(* Logix 5000 project; controller MV vendor 1 type 14 code 217 rev 31.11; software revision 31.00; part 6 of 53 *)
(* tags used below, declared in another part *)
   Alarm_Reset : BOOL;
   Analog_Fault_No : DINT;
   Analog_Simulation_Enabled : BOOL;
   CWD : CHECKWORD_FLAGS;
   Default_Check_Time : DINT;
   FV_YST01_LTX501_AI : PlantItem;   // YST01 LTX501
   FV_YST01_LTX501_AI_RawInput : ALIAS FOR RIO_Rack_2:2:I.Ch2Data;
   FV_YST01_LTX501_ALARM : ALARM_DIGITAL;
   FV_YST01_LTX501_Timer_HiLevel : TIMER;
   FV_YST02_LTX501_AI : PlantItem;   // YST02 LTX501
   FV_YST02_LTX501_AI_RawInput : ALIAS FOR RIO_Rack_2:2:I.Ch3Data;
   FV_YST02_LTX501_ALARM : ALARM_DIGITAL;
   FV_YST02_LTX501_Timer_HiLevel : TIMER;
   FVHRFM03_ALARM : ALARM_DIGITAL;
   FVHRFM03_IP : PlantItem;   // Flow Meter Transmitter
   FVHRFM03_IP_RawInput : ALIAS FOR RIO_Rack_2:16:I.Ch2Data;   // Flow Meter Raw Data
   FVHRLTX02_ALARM : ALARM_DIGITAL;
   FVHRLTX02_IP : PlantItem;   // Effluent Tank Level Transmitter
   FVHRLTX02_IP_Percentage : DINT;
   FVHRLTX02_IP_RawInput : ALIAS FOR RIO_Rack_2:16:I.Ch1Data;   // Effluent Tank Level Transmitter Raw Data
   FVHRLTX02_Timer_HiLevel : TIMER;
   FVHRTM01_IP : PlantItem;   // Turbidty Meter FVHRTM01
   FVHRTM01_IP_RawInput : ALIAS FOR RIO_Rack_2:16:I.Ch0Data;   // Turbidty Meter FVHRTM01 Raw Data
   MC_CH1_CTX1_AI : PlantItem;   // CH1_CTX1
   MC_CH1_CTX1_AI_RawInput : ALIAS FOR RIO_Rack_2:1:I.Ch2Data;   // Real Analog Input , Do Not Use In Code
   MC_CH1_FM_AI : PlantItem;   // CH1_FM
   MC_CH1_FM_AI_RawInput : ALIAS FOR RIO_Rack_2:1:I.Ch4Data;   // Real Analog Input , Do Not Use In Code
   MC_CH1_Log_ID : DINT;
   MC_CH1_PTX_AI : PlantItem;   // CH1_PTX
   MC_CH1_PTX_AI_RawInput : ALIAS FOR RIO_Rack_2:1:I.Ch6Data;   // Real Analog Input , Do Not Use In Code
   MC_CH2_CTX2_AI : PlantItem;   // CH2_CTX2
   MC_CH2_CTX2_AI_RawInput : ALIAS FOR RIO_Rack_2:1:I.Ch3Data;   // Real Analog Input , Do Not Use In Code
   MC_CH2_FM_AI : PlantItem;   // CH2_FM
   MC_CH2_FM_AI_RawInput : ALIAS FOR RIO_Rack_2:1:I.Ch5Data;   // Real Analog Input , Do Not Use In Code
   MC_CH2_Log_ID : DINT;
   MC_CH2_PTX_AI : PlantItem;   // CH2_PTX
   MC_CH2_PTX_AI_RawInput : ALIAS FOR RIO_Rack_2:1:I.Ch7Data;   // Real Analog Input , Do Not Use In Code
   MC_CTX_001_AI : PlantItem;   // CTX_001
   MC_CTX_001_AI_RawInput : ALIAS FOR RIO_Rack_2:1:I.Ch0Data;   // Real Analog Input , Do Not Use In Code
   MC_CTX_002_AI : PlantItem;   // CTX_002
   MC_CTX_002_AI_RawInput : ALIAS FOR RIO_Rack_2:1:I.Ch1Data;   // Real Analog Input , Do Not Use In Code
   MC_N7 : INT[255];   // INTEGER
   MC_P1_SP_AO : PlantItem;   // P1_SP
   MC_P1_SP_AO_RawOutput : ALIAS FOR RIO_Rack_2:3:O.Ch0Data;   // Real Analog Input , Do Not Use In Code
   MC_P2_SP_AO : PlantItem;   // P2_SP
   MC_P2_SP_AO_RawOutput : ALIAS FOR RIO_Rack_2:3:O.Ch1Data;   // Real Analog Input , Do Not Use In Code
   MC_SRV1_Log_ID : DINT;
   MC_SRV2_Log_ID : DINT;
   MC_TTX_001_AI : PlantItem;   // TTX_001
   MC_TTX_001_AI_RawInput : ALIAS FOR RIO_Rack_2:2:I.Ch0Data;   // Real Analog Input , Do Not Use In Code
   MC_TTX_002_AI : PlantItem;   // TTX_002
   MC_TTX_002_AI_RawInput : ALIAS FOR RIO_Rack_2:2:I.Ch1Data;   // Real Analog Input , Do Not Use In Code
   One_Second_One_Scan : ALIAS FOR One_Second_1_scan;
   overrange_RIO_analog_value : REAL;
   underrange_RIO_analog_value : REAL;
   YST_Data : REAL[2];
(* MC_Common, continued *)

ROUTINE MC_A_Events_From_Scada_IDs   (* ladder *)
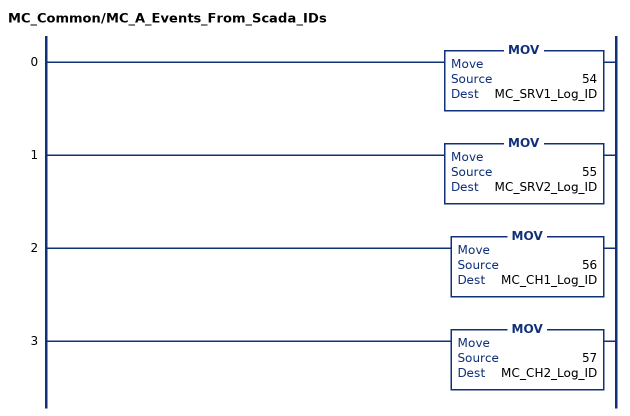
   0: MOV(54,MC_SRV1_Log_ID);
   1: MOV(55,MC_SRV2_Log_ID);
   2: MOV(56,MC_CH1_Log_ID);
   3: MOV(57,MC_CH2_Log_ID);
END_ROUTINE

ROUTINE MC_Analog_Relay_To_NFiles   (* ladder *)
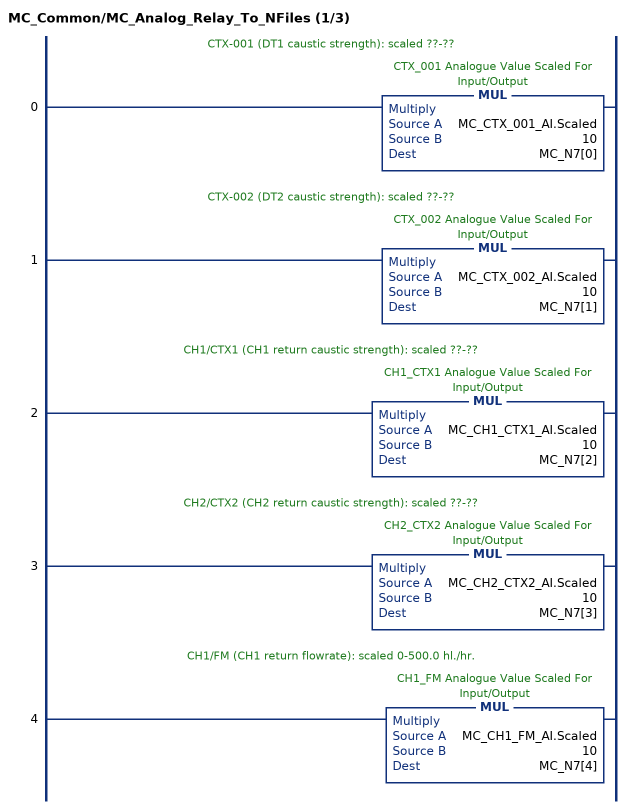
   // CTX-001 (DT1 caustic strength): scaled ??-??
   0: MUL(MC_CTX_001_AI.Scaled,10,MC_N7[0]);
   // CTX-002 (DT2 caustic strength): scaled ??-??
   1: MUL(MC_CTX_002_AI.Scaled,10,MC_N7[1]);
   // CH1/CTX1 (CH1 return caustic strength): scaled ??-??
   2: MUL(MC_CH1_CTX1_AI.Scaled,10,MC_N7[2]);
   // CH2/CTX2 (CH2 return caustic strength): scaled ??-??
   3: MUL(MC_CH2_CTX2_AI.Scaled,10,MC_N7[3]);
   // CH1/FM (CH1 return flowrate): scaled 0-500.0 hl./hr.
   4: MUL(MC_CH1_FM_AI.Scaled,10,MC_N7[4]);
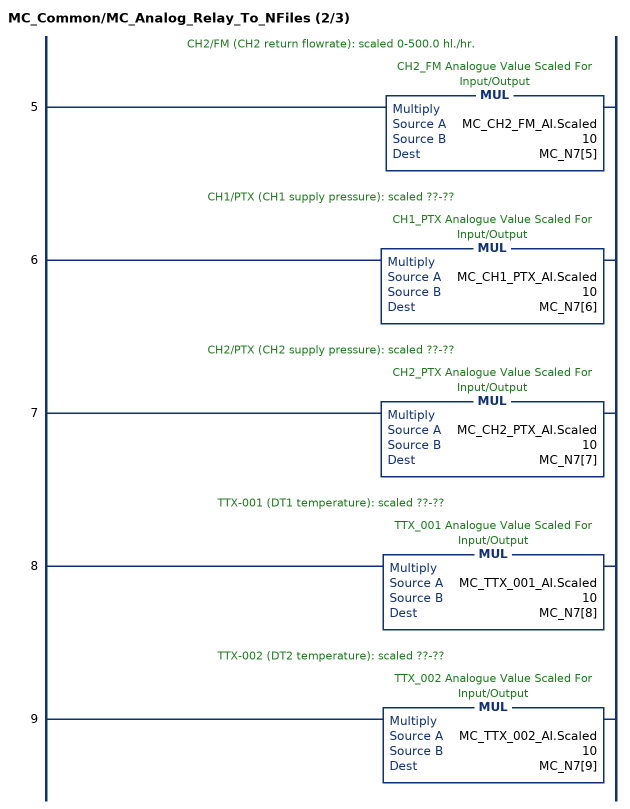
   // CH2/FM (CH2 return flowrate): scaled 0-500.0 hl./hr.
   5: MUL(MC_CH2_FM_AI.Scaled,10,MC_N7[5]);
   // CH1/PTX (CH1 supply pressure): scaled ??-??
   6: MUL(MC_CH1_PTX_AI.Scaled,10,MC_N7[6]);
   // CH2/PTX (CH2 supply pressure): scaled ??-??
   7: MUL(MC_CH2_PTX_AI.Scaled,10,MC_N7[7]);
   // TTX-001 (DT1 temperature): scaled ??-??
   8: MUL(MC_TTX_001_AI.Scaled,10,MC_N7[8]);
   // TTX-002 (DT2 temperature): scaled ??-??
   9: MUL(MC_TTX_002_AI.Scaled,10,MC_N7[9]);
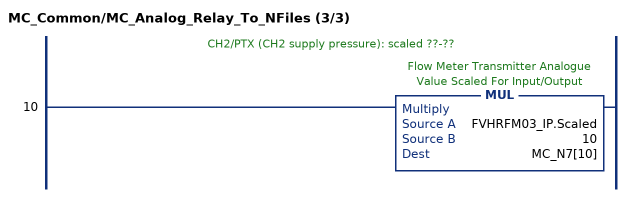
   // CH2/PTX (CH2 supply pressure): scaled ??-??
   10: MUL(FVHRFM03_IP.Scaled,10,MC_N7[10]);
END_ROUTINE

ROUTINE MC_Analogs   (* ladder *)
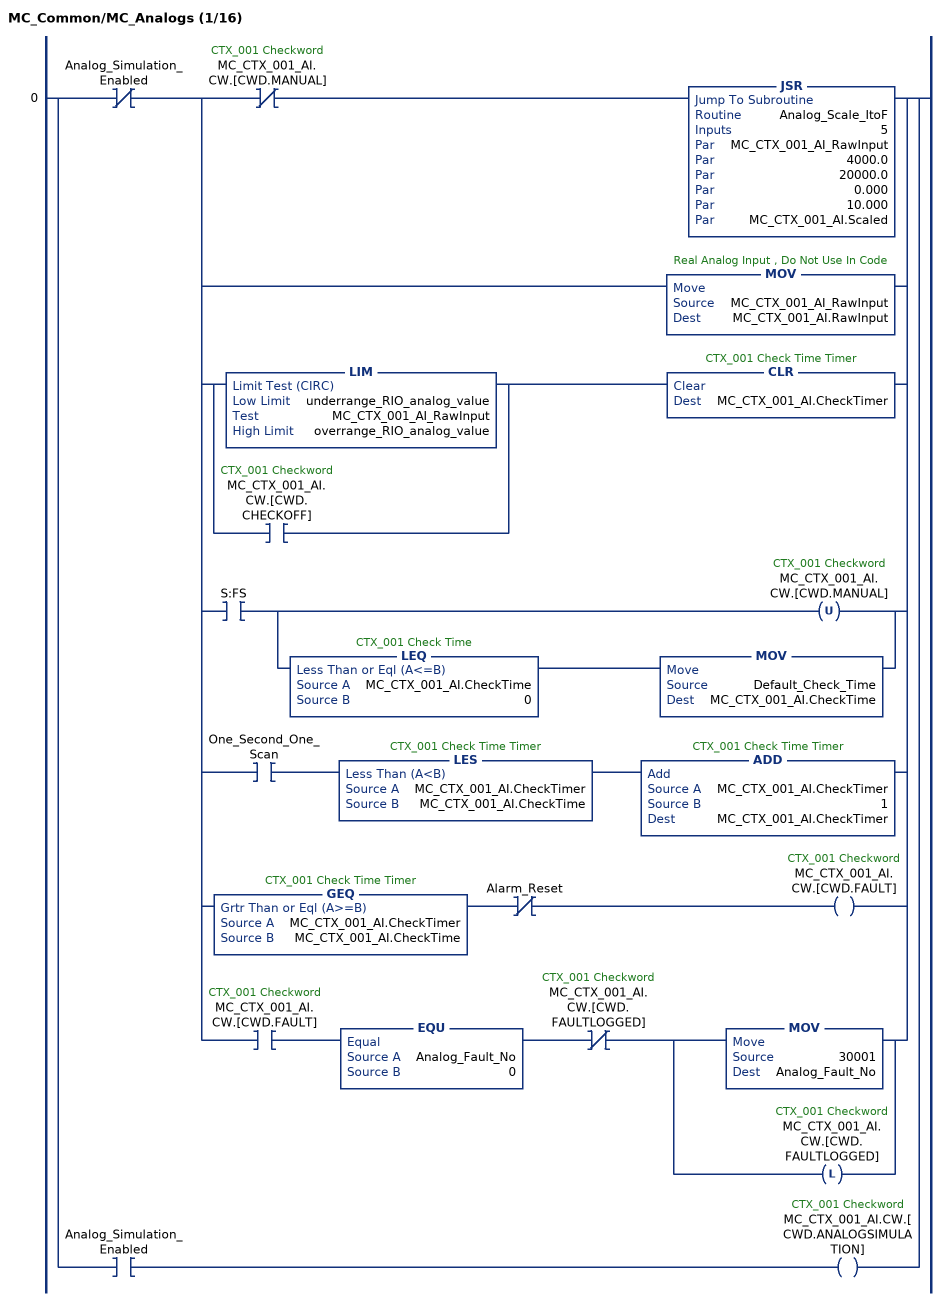
   0: [XIO(Analog_Simulation_Enabled) [XIO(MC_CTX_001_AI.CW.[CWD.MANUAL]) JSR(Analog_Scale_ItoF,5,MC_CTX_001_AI_RawInput,4000.0,20000.0,0.000,10.000,MC_CTX_001_AI.Scaled) ,MOV(MC_CTX_001_AI_RawInput,MC_CTX_001_AI.RawInput) ,[LIM(underrange_RIO_analog_value,MC_CTX_001_AI_RawInput,overrange_RIO_analog_value) ,XIC(MC_CTX_001_AI.CW.[CWD.CHECKOFF]) ] CLR(MC_CTX_001_AI.CheckTimer) ,XIC(S:FS) [OTU(MC_CTX_001_AI.CW.[CWD.MANUAL]) ,LEQ(MC_CTX_001_AI.CheckTime,0) MOV(Default_Check_Time,MC_CTX_001_AI.CheckTime) ] ,XIC(One_Second_One_Scan) LES(MC_CTX_001_AI.CheckTimer,MC_CTX_001_AI.CheckTime) ADD(MC_CTX_001_AI.CheckTimer,1,MC_CTX_001_AI.CheckTimer) ,GEQ(MC_CTX_001_AI.CheckTimer,MC_CTX_001_AI.CheckTime) XIO(Alarm_Reset) OTE(MC_CTX_001_AI.CW.[CWD.FAULT]) ,XIC(MC_CTX_001_AI.CW.[CWD.FAULT]) EQU(Analog_Fault_No,0) XIO(MC_CTX_001_AI.CW.[CWD.FAULTLOGGED]) [MOV(30001,Analog_Fault_No) ,OTL(MC_CTX_001_AI.CW.[CWD.FAULTLOGGED]) ] ] ,XIC(Analog_Simulation_Enabled) OTE(MC_CTX_001_AI.CW.[CWD.ANALOGSIMULATION]) ];
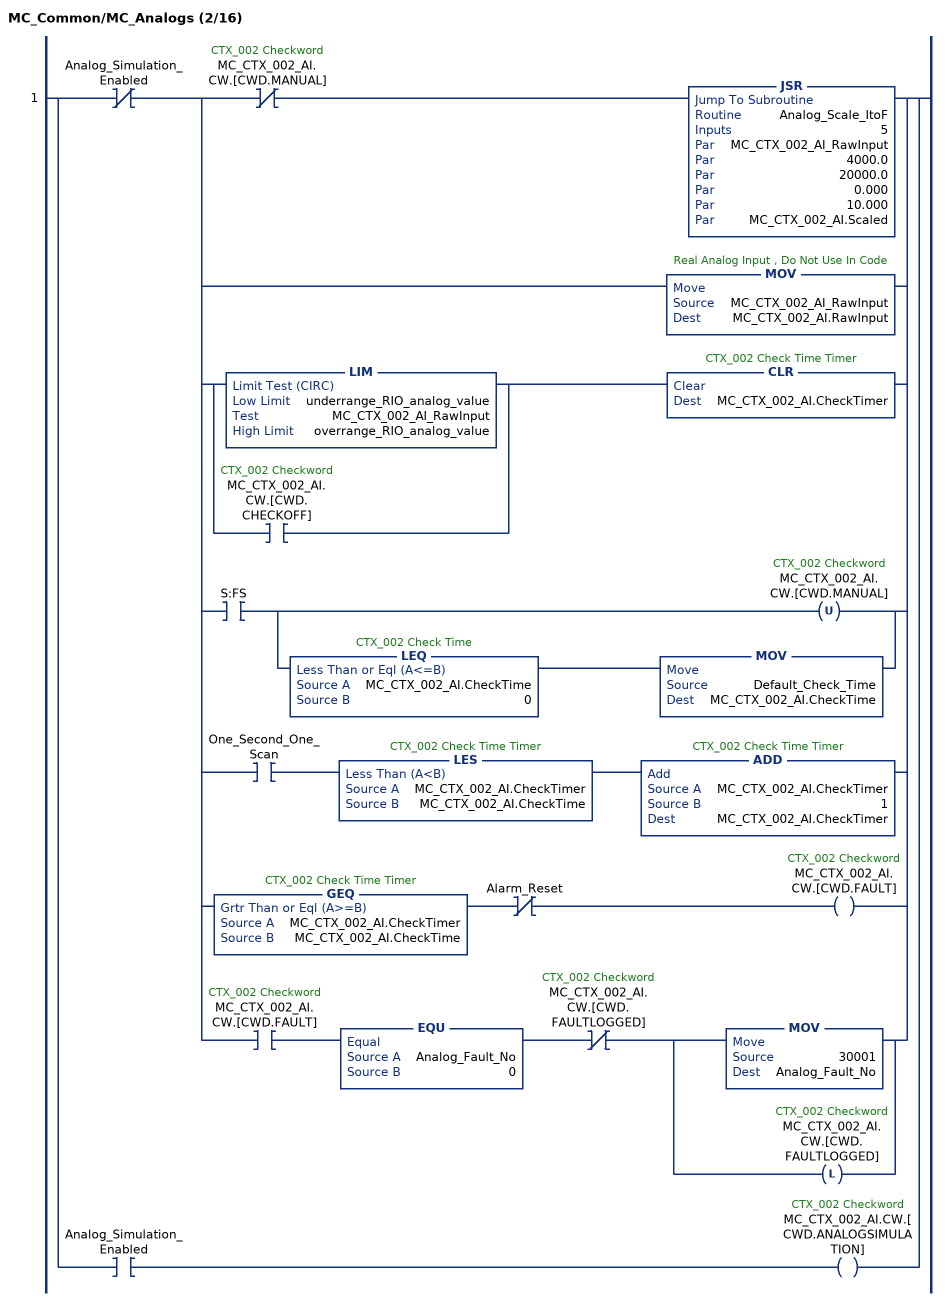
   1: [XIO(Analog_Simulation_Enabled) [XIO(MC_CTX_002_AI.CW.[CWD.MANUAL]) JSR(Analog_Scale_ItoF,5,MC_CTX_002_AI_RawInput,4000.0,20000.0,0.000,10.000,MC_CTX_002_AI.Scaled) ,MOV(MC_CTX_002_AI_RawInput,MC_CTX_002_AI.RawInput) ,[LIM(underrange_RIO_analog_value,MC_CTX_002_AI_RawInput,overrange_RIO_analog_value) ,XIC(MC_CTX_002_AI.CW.[CWD.CHECKOFF]) ] CLR(MC_CTX_002_AI.CheckTimer) ,XIC(S:FS) [OTU(MC_CTX_002_AI.CW.[CWD.MANUAL]) ,LEQ(MC_CTX_002_AI.CheckTime,0) MOV(Default_Check_Time,MC_CTX_002_AI.CheckTime) ] ,XIC(One_Second_One_Scan) LES(MC_CTX_002_AI.CheckTimer,MC_CTX_002_AI.CheckTime) ADD(MC_CTX_002_AI.CheckTimer,1,MC_CTX_002_AI.CheckTimer) ,GEQ(MC_CTX_002_AI.CheckTimer,MC_CTX_002_AI.CheckTime) XIO(Alarm_Reset) OTE(MC_CTX_002_AI.CW.[CWD.FAULT]) ,XIC(MC_CTX_002_AI.CW.[CWD.FAULT]) EQU(Analog_Fault_No,0) XIO(MC_CTX_002_AI.CW.[CWD.FAULTLOGGED]) [MOV(30001,Analog_Fault_No) ,OTL(MC_CTX_002_AI.CW.[CWD.FAULTLOGGED]) ] ] ,XIC(Analog_Simulation_Enabled) OTE(MC_CTX_002_AI.CW.[CWD.ANALOGSIMULATION]) ];
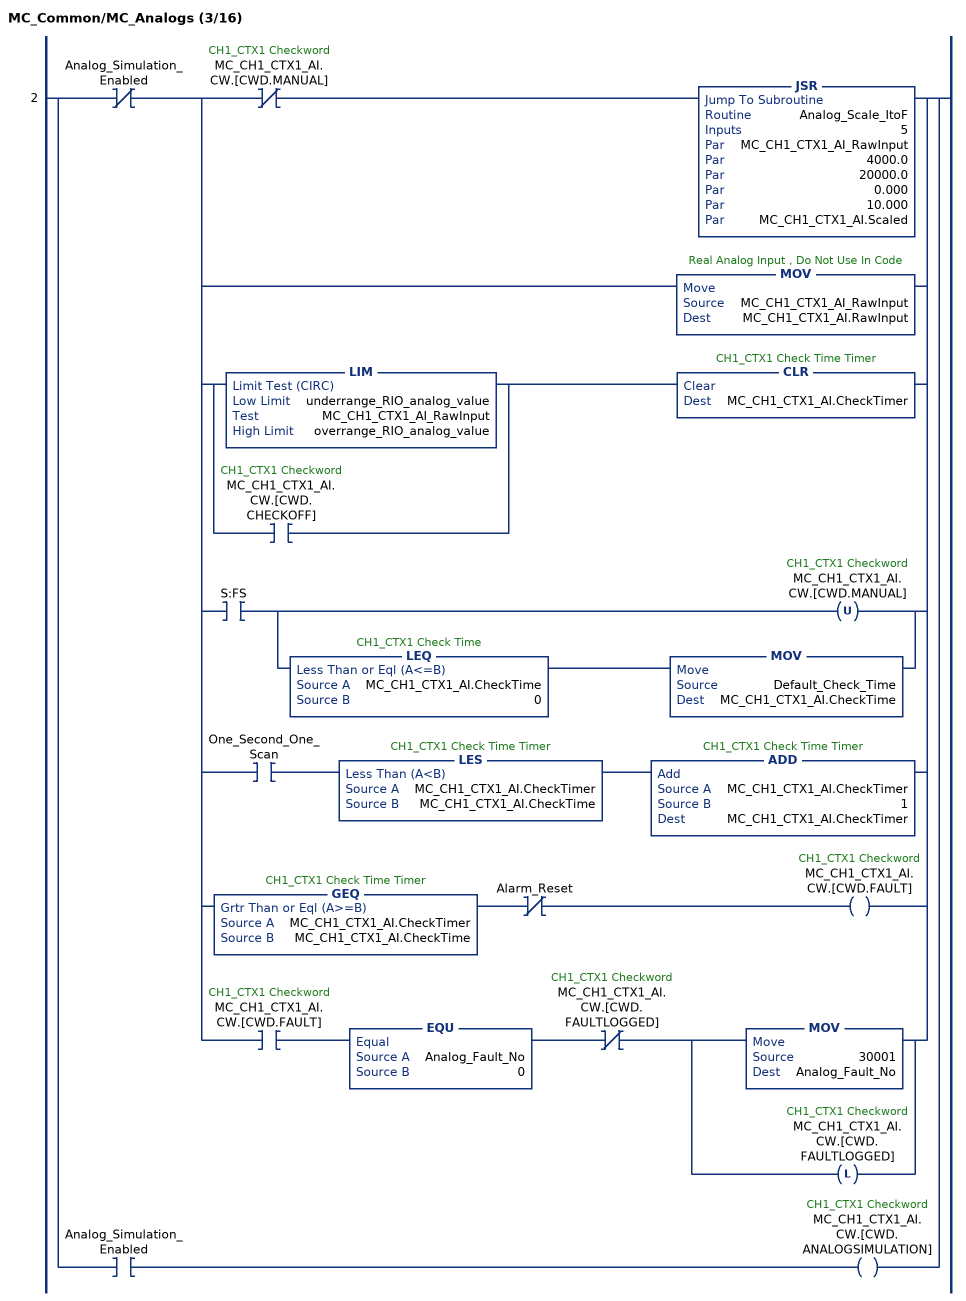
   2: [XIO(Analog_Simulation_Enabled) [XIO(MC_CH1_CTX1_AI.CW.[CWD.MANUAL]) JSR(Analog_Scale_ItoF,5,MC_CH1_CTX1_AI_RawInput,4000.0,20000.0,0.000,10.000,MC_CH1_CTX1_AI.Scaled) ,MOV(MC_CH1_CTX1_AI_RawInput,MC_CH1_CTX1_AI.RawInput) ,[LIM(underrange_RIO_analog_value,MC_CH1_CTX1_AI_RawInput,overrange_RIO_analog_value) ,XIC(MC_CH1_CTX1_AI.CW.[CWD.CHECKOFF]) ] CLR(MC_CH1_CTX1_AI.CheckTimer) ,XIC(S:FS) [OTU(MC_CH1_CTX1_AI.CW.[CWD.MANUAL]) ,LEQ(MC_CH1_CTX1_AI.CheckTime,0) MOV(Default_Check_Time,MC_CH1_CTX1_AI.CheckTime) ] ,XIC(One_Second_One_Scan) LES(MC_CH1_CTX1_AI.CheckTimer,MC_CH1_CTX1_AI.CheckTime) ADD(MC_CH1_CTX1_AI.CheckTimer,1,MC_CH1_CTX1_AI.CheckTimer) ,GEQ(MC_CH1_CTX1_AI.CheckTimer,MC_CH1_CTX1_AI.CheckTime) XIO(Alarm_Reset) OTE(MC_CH1_CTX1_AI.CW.[CWD.FAULT]) ,XIC(MC_CH1_CTX1_AI.CW.[CWD.FAULT]) EQU(Analog_Fault_No,0) XIO(MC_CH1_CTX1_AI.CW.[CWD.FAULTLOGGED]) [MOV(30001,Analog_Fault_No) ,OTL(MC_CH1_CTX1_AI.CW.[CWD.FAULTLOGGED]) ] ] ,XIC(Analog_Simulation_Enabled) OTE(MC_CH1_CTX1_AI.CW.[CWD.ANALOGSIMULATION]) ];
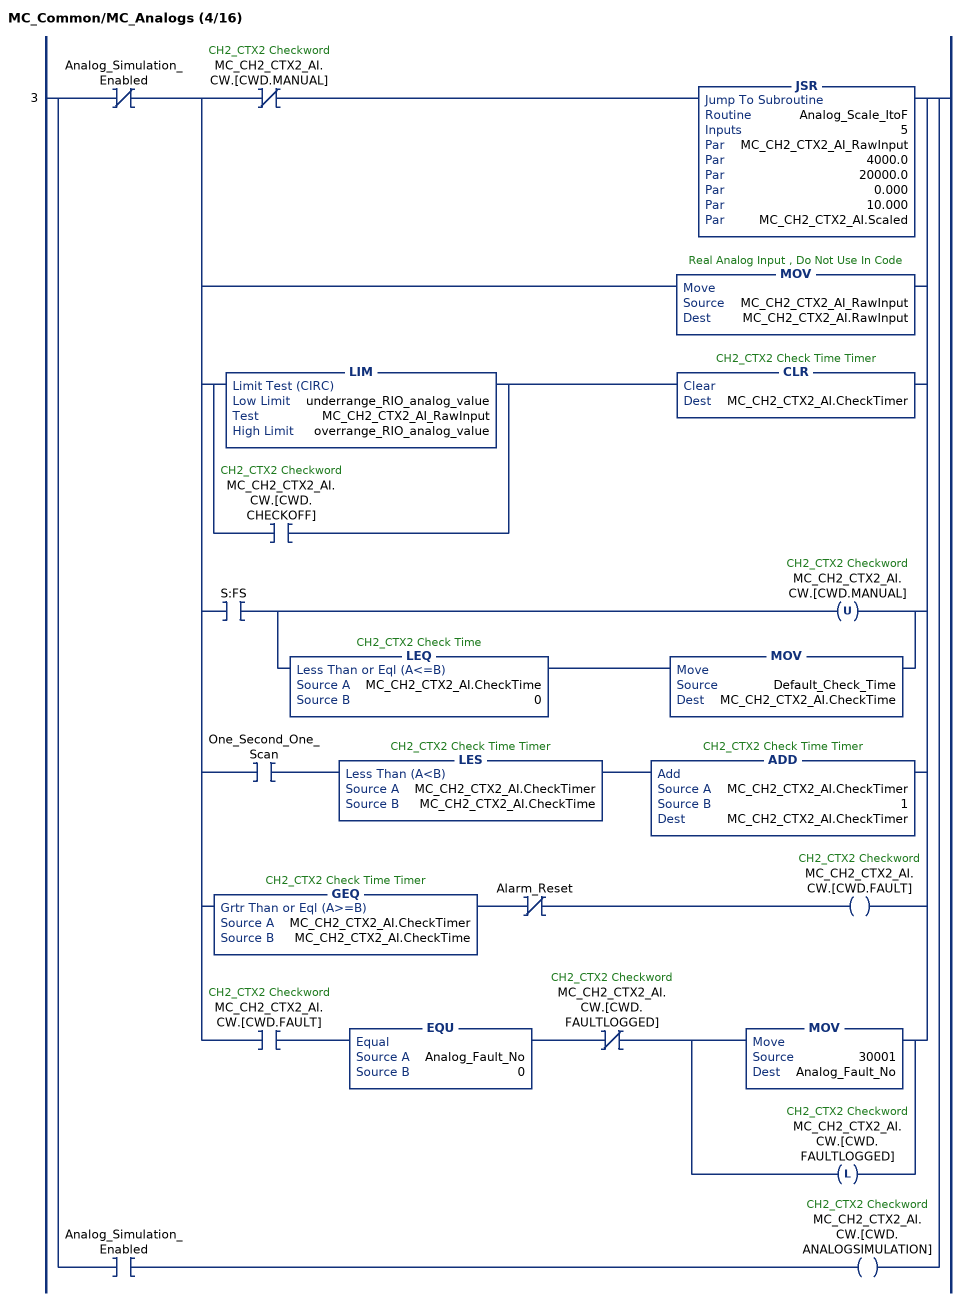
   3: [XIO(Analog_Simulation_Enabled) [XIO(MC_CH2_CTX2_AI.CW.[CWD.MANUAL]) JSR(Analog_Scale_ItoF,5,MC_CH2_CTX2_AI_RawInput,4000.0,20000.0,0.000,10.000,MC_CH2_CTX2_AI.Scaled) ,MOV(MC_CH2_CTX2_AI_RawInput,MC_CH2_CTX2_AI.RawInput) ,[LIM(underrange_RIO_analog_value,MC_CH2_CTX2_AI_RawInput,overrange_RIO_analog_value) ,XIC(MC_CH2_CTX2_AI.CW.[CWD.CHECKOFF]) ] CLR(MC_CH2_CTX2_AI.CheckTimer) ,XIC(S:FS) [OTU(MC_CH2_CTX2_AI.CW.[CWD.MANUAL]) ,LEQ(MC_CH2_CTX2_AI.CheckTime,0) MOV(Default_Check_Time,MC_CH2_CTX2_AI.CheckTime) ] ,XIC(One_Second_One_Scan) LES(MC_CH2_CTX2_AI.CheckTimer,MC_CH2_CTX2_AI.CheckTime) ADD(MC_CH2_CTX2_AI.CheckTimer,1,MC_CH2_CTX2_AI.CheckTimer) ,GEQ(MC_CH2_CTX2_AI.CheckTimer,MC_CH2_CTX2_AI.CheckTime) XIO(Alarm_Reset) OTE(MC_CH2_CTX2_AI.CW.[CWD.FAULT]) ,XIC(MC_CH2_CTX2_AI.CW.[CWD.FAULT]) EQU(Analog_Fault_No,0) XIO(MC_CH2_CTX2_AI.CW.[CWD.FAULTLOGGED]) [MOV(30001,Analog_Fault_No) ,OTL(MC_CH2_CTX2_AI.CW.[CWD.FAULTLOGGED]) ] ] ,XIC(Analog_Simulation_Enabled) OTE(MC_CH2_CTX2_AI.CW.[CWD.ANALOGSIMULATION]) ];
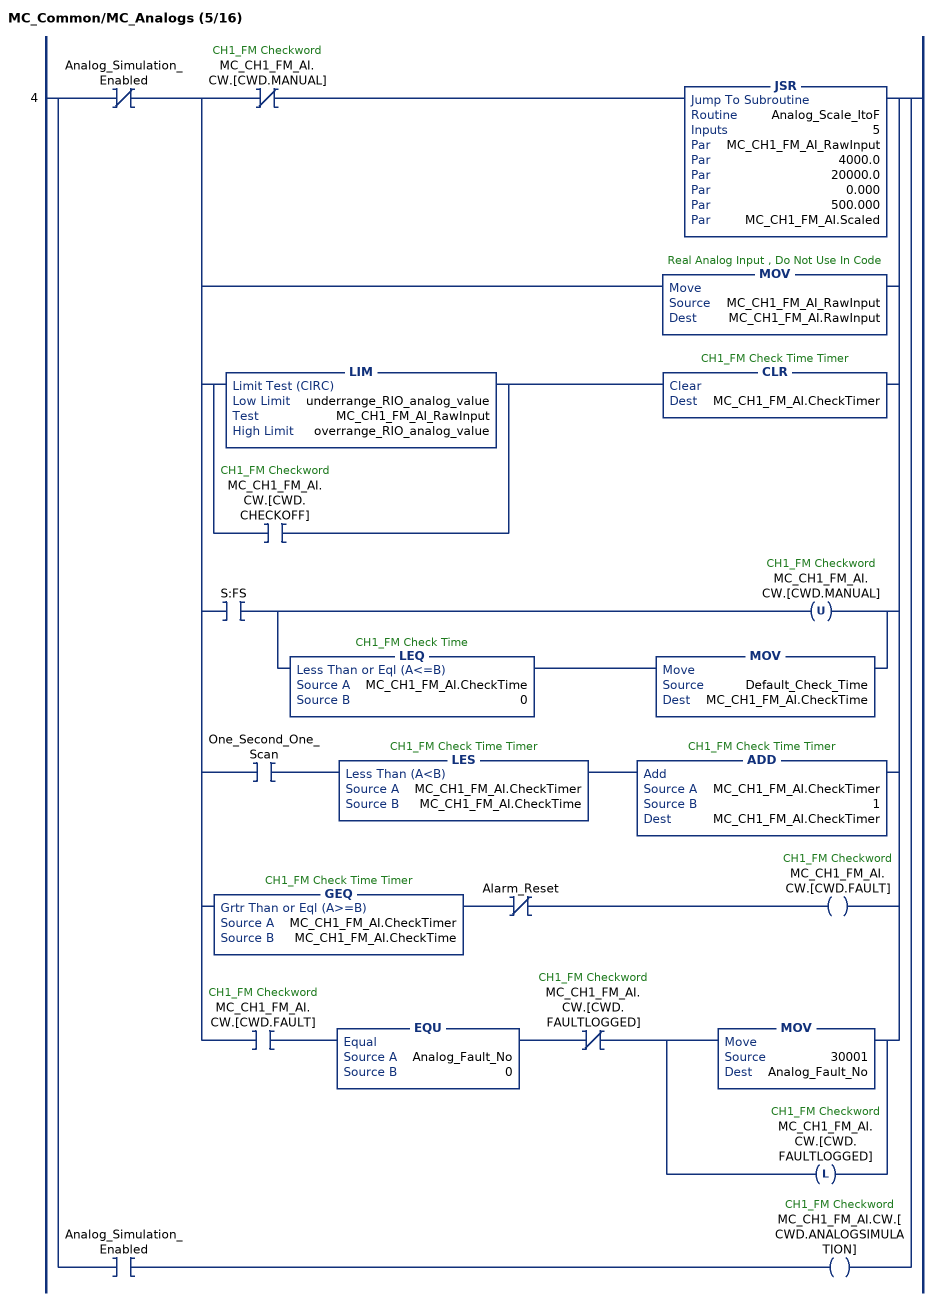
   4: [XIO(Analog_Simulation_Enabled) [XIO(MC_CH1_FM_AI.CW.[CWD.MANUAL]) JSR(Analog_Scale_ItoF,5,MC_CH1_FM_AI_RawInput,4000.0,20000.0,0.000,500.000,MC_CH1_FM_AI.Scaled) ,MOV(MC_CH1_FM_AI_RawInput,MC_CH1_FM_AI.RawInput) ,[LIM(underrange_RIO_analog_value,MC_CH1_FM_AI_RawInput,overrange_RIO_analog_value) ,XIC(MC_CH1_FM_AI.CW.[CWD.CHECKOFF]) ] CLR(MC_CH1_FM_AI.CheckTimer) ,XIC(S:FS) [OTU(MC_CH1_FM_AI.CW.[CWD.MANUAL]) ,LEQ(MC_CH1_FM_AI.CheckTime,0) MOV(Default_Check_Time,MC_CH1_FM_AI.CheckTime) ] ,XIC(One_Second_One_Scan) LES(MC_CH1_FM_AI.CheckTimer,MC_CH1_FM_AI.CheckTime) ADD(MC_CH1_FM_AI.CheckTimer,1,MC_CH1_FM_AI.CheckTimer) ,GEQ(MC_CH1_FM_AI.CheckTimer,MC_CH1_FM_AI.CheckTime) XIO(Alarm_Reset) OTE(MC_CH1_FM_AI.CW.[CWD.FAULT]) ,XIC(MC_CH1_FM_AI.CW.[CWD.FAULT]) EQU(Analog_Fault_No,0) XIO(MC_CH1_FM_AI.CW.[CWD.FAULTLOGGED]) [MOV(30001,Analog_Fault_No) ,OTL(MC_CH1_FM_AI.CW.[CWD.FAULTLOGGED]) ] ] ,XIC(Analog_Simulation_Enabled) OTE(MC_CH1_FM_AI.CW.[CWD.ANALOGSIMULATION]) ];
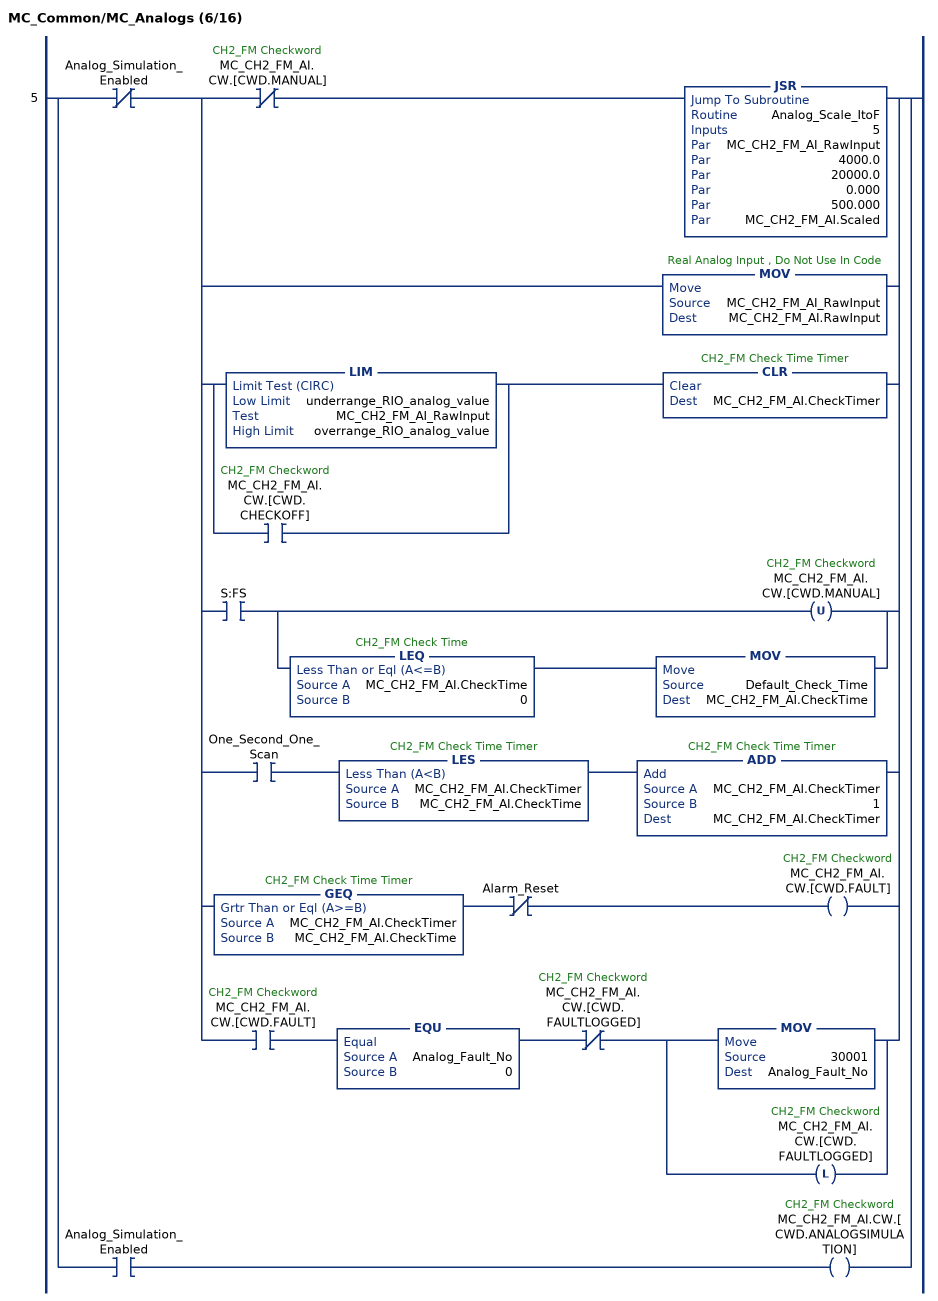
   5: [XIO(Analog_Simulation_Enabled) [XIO(MC_CH2_FM_AI.CW.[CWD.MANUAL]) JSR(Analog_Scale_ItoF,5,MC_CH2_FM_AI_RawInput,4000.0,20000.0,0.000,500.000,MC_CH2_FM_AI.Scaled) ,MOV(MC_CH2_FM_AI_RawInput,MC_CH2_FM_AI.RawInput) ,[LIM(underrange_RIO_analog_value,MC_CH2_FM_AI_RawInput,overrange_RIO_analog_value) ,XIC(MC_CH2_FM_AI.CW.[CWD.CHECKOFF]) ] CLR(MC_CH2_FM_AI.CheckTimer) ,XIC(S:FS) [OTU(MC_CH2_FM_AI.CW.[CWD.MANUAL]) ,LEQ(MC_CH2_FM_AI.CheckTime,0) MOV(Default_Check_Time,MC_CH2_FM_AI.CheckTime) ] ,XIC(One_Second_One_Scan) LES(MC_CH2_FM_AI.CheckTimer,MC_CH2_FM_AI.CheckTime) ADD(MC_CH2_FM_AI.CheckTimer,1,MC_CH2_FM_AI.CheckTimer) ,GEQ(MC_CH2_FM_AI.CheckTimer,MC_CH2_FM_AI.CheckTime) XIO(Alarm_Reset) OTE(MC_CH2_FM_AI.CW.[CWD.FAULT]) ,XIC(MC_CH2_FM_AI.CW.[CWD.FAULT]) EQU(Analog_Fault_No,0) XIO(MC_CH2_FM_AI.CW.[CWD.FAULTLOGGED]) [MOV(30001,Analog_Fault_No) ,OTL(MC_CH2_FM_AI.CW.[CWD.FAULTLOGGED]) ] ] ,XIC(Analog_Simulation_Enabled) OTE(MC_CH2_FM_AI.CW.[CWD.ANALOGSIMULATION]) ];